   // Erhöhen des Gesammtverbrauches und des Gesamtzählers:
   // 
   "DB_Zaehler_Schicht_aktuell".Gesamt.Anzahl := "DB_Zaehler_Schicht_aktuell".Gesamt.Anzahl + 1;
   (* classic code: "DB_Zaehler_Schicht_aktuell".Gesamt.Verbrauch_K1 :=  "DB_Zaehler_Schicht_aktuell".Gesamt.Verbrauch_K1 + "DB919_ShotResultMach".ShotResult_Ma[0].Component.Comp[1].MaterialConsumption / 1000.0;*)
   "DB_Zaehler_Schicht_aktuell".Gesamt.Verbrauch_K1 :=  "DB_Zaehler_Schicht_aktuell".Gesamt.Verbrauch_K1 + "DB919_ShotResultMach".ShotResult_Ma[0].Component.Comp[1].MaterialConsumption / REAL#1000.0;
   (* classic code: "DB_Zaehler_Schicht_aktuell".Gesamt.Verbrauch_K2 :=  "DB_Zaehler_Schicht_aktuell".Gesamt.Verbrauch_K2 + "DB919_ShotResultMach".ShotResult_Ma[0].Component.Comp[2].MaterialConsumption / 1000.0;*)
   "DB_Zaehler_Schicht_aktuell".Gesamt.Verbrauch_K2 :=  "DB_Zaehler_Schicht_aktuell".Gesamt.Verbrauch_K2 + "DB919_ShotResultMach".ShotResult_Ma[0].Component.Comp[2].MaterialConsumption / REAL#1000.0;
   (* classic code: "DB_Zaehler_Schicht_aktuell".Gesamt.Verbrauch_K3 :=  "DB_Zaehler_Schicht_aktuell".Gesamt.Verbrauch_K3 + "DB919_ShotResultMach".ShotResult_Ma[0].Component.Comp[3].MaterialConsumption / 1000.0;*)
   "DB_Zaehler_Schicht_aktuell".Gesamt.Verbrauch_K3 :=  "DB_Zaehler_Schicht_aktuell".Gesamt.Verbrauch_K3 + "DB919_ShotResultMach".ShotResult_Ma[0].Component.Comp[3].MaterialConsumption / REAL#1000.0;
   (* classic code: "DB_Zaehler_Schicht_aktuell".Gesamt.Verbrauch_K4 :=  "DB_Zaehler_Schicht_aktuell".Gesamt.Verbrauch_K4 + "DB919_ShotResultMach".ShotResult_Ma[0].Component.Comp[4].MaterialConsumption / 1000.0;*)
   "DB_Zaehler_Schicht_aktuell".Gesamt.Verbrauch_K4 :=  "DB_Zaehler_Schicht_aktuell".Gesamt.Verbrauch_K4 + "DB919_ShotResultMach".ShotResult_Ma[0].Component.Comp[4].MaterialConsumption / REAL#1000.0;
   (* classic code: "DB_Zaehler_Schicht_aktuell".Gesamt.Verbrauch_K5 :=  "DB_Zaehler_Schicht_aktuell".Gesamt.Verbrauch_K5 + "DB919_ShotResultMach".ShotResult_Ma[0].Component.Comp[5].MaterialConsumption / 1000.0;*)
   "DB_Zaehler_Schicht_aktuell".Gesamt.Verbrauch_K5 :=  "DB_Zaehler_Schicht_aktuell".Gesamt.Verbrauch_K5 + "DB919_ShotResultMach".ShotResult_Ma[0].Component.Comp[5].MaterialConsumption / REAL#1000.0;
   (* classic code: "DB_Zaehler_Schicht_aktuell".Gesamt.Verbrauch_K6 :=  "DB_Zaehler_Schicht_aktuell".Gesamt.Verbrauch_K6 + "DB919_ShotResultMach".ShotResult_Ma[0].Component.Comp[6].MaterialConsumption / 1000.0;*)
   "DB_Zaehler_Schicht_aktuell".Gesamt.Verbrauch_K6 :=  "DB_Zaehler_Schicht_aktuell".Gesamt.Verbrauch_K6 + "DB919_ShotResultMach".ShotResult_Ma[0].Component.Comp[6].MaterialConsumption / REAL#1000.0;
   (* classic code: "DB_Zaehler_Schicht_aktuell".Gesamt.Verbrauch_K7 :=  "DB_Zaehler_Schicht_aktuell".Gesamt.Verbrauch_K7 + "DB919_ShotResultMach".ShotResult_Ma[0].Component.Comp[7].MaterialConsumption / 1000.0;*)
   "DB_Zaehler_Schicht_aktuell".Gesamt.Verbrauch_K7 :=  "DB_Zaehler_Schicht_aktuell".Gesamt.Verbrauch_K7 + "DB919_ShotResultMach".ShotResult_Ma[0].Component.Comp[7].MaterialConsumption / REAL#1000.0;
   (* classic code: "DB_Zaehler_Schicht_aktuell".Gesamt.Verbrauch_K8 :=  "DB_Zaehler_Schicht_aktuell".Gesamt.Verbrauch_K8 + "DB919_ShotResultMach".ShotResult_Ma[0].Component.Comp[8].MaterialConsumption / 1000.0;*)
   "DB_Zaehler_Schicht_aktuell".Gesamt.Verbrauch_K8 :=  "DB_Zaehler_Schicht_aktuell".Gesamt.Verbrauch_K8 + "DB919_ShotResultMach".ShotResult_Ma[0].Component.Comp[8].MaterialConsumption / REAL#1000.0;

   // Erhöhen des im Programm eingetragenen Schußzählers:
   // 
   // Benötigte Variablen:
   // der aktuelle Teiezähler: "DB919_ShotResultMach".ShotResult_Ma[0].General.PartID
   // 
   IF "DB919_ShotResultMach".ShotResult_Ma[0].General.PartID > 0 THEN
     #i := "DB919_ShotResultMach".ShotResult_Ma[0].General.PartID;
     "DB_Zaehler_Schicht_aktuell".Counter[#i].Anzahl := "DB_Zaehler_Schicht_aktuell".Counter[#i].Anzahl + 1;
     (* classic code: "DB_Zaehler_Schicht_aktuell".Counter[#i].Verbrauch_K1 := "DB_Zaehler_Schicht_aktuell".Counter[#i].Verbrauch_K1 + "DB919_ShotResultMach".ShotResult_Ma[0].Component.Comp[1].MaterialConsumption / 1000.0;*)
     "DB_Zaehler_Schicht_aktuell".Counter[#i].Verbrauch_K1 := "DB_Zaehler_Schicht_aktuell".Counter[#i].Verbrauch_K1 + "DB919_ShotResultMach".ShotResult_Ma[0].Component.Comp[1].MaterialConsumption / REAL#1000.0;
     (* classic code: "DB_Zaehler_Schicht_aktuell".Counter[#i].Verbrauch_K2 := "DB_Zaehler_Schicht_aktuell".Counter[#i].Verbrauch_K2 + "DB919_ShotResultMach".ShotResult_Ma[0].Component.Comp[2].MaterialConsumption / 1000.0;*)
     "DB_Zaehler_Schicht_aktuell".Counter[#i].Verbrauch_K2 := "DB_Zaehler_Schicht_aktuell".Counter[#i].Verbrauch_K2 + "DB919_ShotResultMach".ShotResult_Ma[0].Component.Comp[2].MaterialConsumption / REAL#1000.0;
     (* classic code: "DB_Zaehler_Schicht_aktuell".Counter[#i].Verbrauch_K3 := "DB_Zaehler_Schicht_aktuell".Counter[#i].Verbrauch_K3 + "DB919_ShotResultMach".ShotResult_Ma[0].Component.Comp[3].MaterialConsumption / 1000.0;*)
     "DB_Zaehler_Schicht_aktuell".Counter[#i].Verbrauch_K3 := "DB_Zaehler_Schicht_aktuell".Counter[#i].Verbrauch_K3 + "DB919_ShotResultMach".ShotResult_Ma[0].Component.Comp[3].MaterialConsumption / REAL#1000.0;
     (* classic code: "DB_Zaehler_Schicht_aktuell".Counter[#i].Verbrauch_K4 := "DB_Zaehler_Schicht_aktuell".Counter[#i].Verbrauch_K4 + "DB919_ShotResultMach".ShotResult_Ma[0].Component.Comp[4].MaterialConsumption / 1000.0;*)
     "DB_Zaehler_Schicht_aktuell".Counter[#i].Verbrauch_K4 := "DB_Zaehler_Schicht_aktuell".Counter[#i].Verbrauch_K4 + "DB919_ShotResultMach".ShotResult_Ma[0].Component.Comp[4].MaterialConsumption / REAL#1000.0;
     (* classic code: "DB_Zaehler_Schicht_aktuell".Counter[#i].Verbrauch_K5 := "DB_Zaehler_Schicht_aktuell".Counter[#i].Verbrauch_K5 + "DB919_ShotResultMach".ShotResult_Ma[0].Component.Comp[5].MaterialConsumption / 1000.0;*)
     "DB_Zaehler_Schicht_aktuell".Counter[#i].Verbrauch_K5 := "DB_Zaehler_Schicht_aktuell".Counter[#i].Verbrauch_K5 + "DB919_ShotResultMach".ShotResult_Ma[0].Component.Comp[5].MaterialConsumption / REAL#1000.0;
     (* classic code: "DB_Zaehler_Schicht_aktuell".Counter[#i].Verbrauch_K6 := "DB_Zaehler_Schicht_aktuell".Counter[#i].Verbrauch_K6 + "DB919_ShotResultMach".ShotResult_Ma[0].Component.Comp[6].MaterialConsumption / 1000.0;*)
     "DB_Zaehler_Schicht_aktuell".Counter[#i].Verbrauch_K6 := "DB_Zaehler_Schicht_aktuell".Counter[#i].Verbrauch_K6 + "DB919_ShotResultMach".ShotResult_Ma[0].Component.Comp[6].MaterialConsumption / REAL#1000.0;
     (* classic code: "DB_Zaehler_Schicht_aktuell".Counter[#i].Verbrauch_K7 := "DB_Zaehler_Schicht_aktuell".Counter[#i].Verbrauch_K7 + "DB919_ShotResultMach".ShotResult_Ma[0].Component.Comp[7].MaterialConsumption / 1000.0;*)
     "DB_Zaehler_Schicht_aktuell".Counter[#i].Verbrauch_K7 := "DB_Zaehler_Schicht_aktuell".Counter[#i].Verbrauch_K7 + "DB919_ShotResultMach".ShotResult_Ma[0].Component.Comp[7].MaterialConsumption / REAL#1000.0;
     (* classic code: "DB_Zaehler_Schicht_aktuell".Counter[#i].Verbrauch_K8 := "DB_Zaehler_Schicht_aktuell".Counter[#i].Verbrauch_K8 + "DB919_ShotResultMach".ShotResult_Ma[0].Component.Comp[8].MaterialConsumption / 1000.0;*)
     "DB_Zaehler_Schicht_aktuell".Counter[#i].Verbrauch_K8 := "DB_Zaehler_Schicht_aktuell".Counter[#i].Verbrauch_K8 + "DB919_ShotResultMach".ShotResult_Ma[0].Component.Comp[8].MaterialConsumption / REAL#1000.0;
   END_IF;
END_FUNCTION

FUNCTION "PartCounterView" : Void   // FC5002, SCL
{ S7_Optimized_Access := 'FALSE' }
VERSION : 0.1
   VAR_TEMP
      i : Int;
      CounterStartNumber : Int;
   END_VAR
BEGIN
   #CounterStartNumber := "DB_Zaehler_Anzeige".ReadWriteDeviceNo;

   IF "DB_Zaehler_Anzeige".Read THEN
     IF "DB_Zaehler_Anzeige".ViewPreShift = 0 THEN
       FOR #i := 1 TO 10 DO
         "DB_Zaehler_Anzeige".Counter[#i] :="DB_Zaehler_Schicht_aktuell".Counter[#CounterStartNumber];
         #CounterStartNumber := #CounterStartNumber +1;
       END_FOR;
       "DB_Zaehler_Anzeige".Gesamt := "DB_Zaehler_Schicht_aktuell".Gesamt;
       "DB_Zaehler_Anzeige".MH_Counter_ActualShift := "DB_Zaehler_Schicht_aktuell".MH_Counter;
     ELSE
       FOR #i := 1 TO 10 DO
         "DB_Zaehler_Anzeige".Counter[#i] :="DB_Zaehler_Schicht_Vorherige".Counter[#CounterStartNumber];
         #CounterStartNumber := #CounterStartNumber +1;
       END_FOR;
       "DB_Zaehler_Anzeige".Gesamt := "DB_Zaehler_Schicht_Vorherige".Gesamt;
       "DB_Zaehler_Anzeige".MH_Counter_ActualShift := "DB_Zaehler_Schicht_Vorherige".MH_Counter;
     END_IF;

     FOR #i := 1 TO 16 DO
       "DB_Zaehler_Anzeige".MH_Counter_ActualShift[#i] := "DB_Zaehler_Schicht_aktuell".MH_Counter[#i];
       "DB_Zaehler_Anzeige".MH_Counter_PreShift[#i] :=  "DB_Zaehler_Schicht_Vorherige".MH_Counter[#i];
     END_FOR;

   END_IF;

   "DB_Zaehler_Anzeige".Read := false;
END_FUNCTION

FUNCTION "PartCounterCopy" : Void   // FC5003, SCL
{ S7_Optimized_Access := 'FALSE' }
VERSION : 0.1
   VAR_TEMP
      i : Int;
   END_VAR
BEGIN
   // 
   // Shift the part counter at the begining of a new shift!
   // 
   "DB_Zaehler_Schicht_Vorherige".Gesamt := "DB_Zaehler_Schicht_aktuell".Gesamt;
   "DB_Zaehler_Schicht_Vorherige".Counter := "DB_Zaehler_Schicht_aktuell".Counter;
   "DB_Zaehler_Schicht_Vorherige".MH_Counter := "DB_Zaehler_Schicht_aktuell".MH_Counter;

   // Reset the amount of Counts and weight
   // 
   "DB_Zaehler_Schicht_aktuell".Gesamt.Anzahl := 0;
   (* classic code: "DB_Zaehler_Schicht_aktuell".Gesamt.Verbrauch_K1 := 0.0;*)
   "DB_Zaehler_Schicht_aktuell".Gesamt.Verbrauch_K1 := REAL#0.0;
   (* classic code: "DB_Zaehler_Schicht_aktuell".Gesamt.Verbrauch_K2 := 0.0;*)
   "DB_Zaehler_Schicht_aktuell".Gesamt.Verbrauch_K2 := REAL#0.0;
   (* classic code: "DB_Zaehler_Schicht_aktuell".Gesamt.Verbrauch_K3 := 0.0;*)
   "DB_Zaehler_Schicht_aktuell".Gesamt.Verbrauch_K3 := REAL#0.0;
   (* classic code: "DB_Zaehler_Schicht_aktuell".Gesamt.Verbrauch_K4 := 0.0;*)
   "DB_Zaehler_Schicht_aktuell".Gesamt.Verbrauch_K4 := REAL#0.0;
   (* classic code: "DB_Zaehler_Schicht_aktuell".Gesamt.Verbrauch_K5 := 0.0;*)
   "DB_Zaehler_Schicht_aktuell".Gesamt.Verbrauch_K5 := REAL#0.0;
   (* classic code: "DB_Zaehler_Schicht_aktuell".Gesamt.Verbrauch_K6 := 0.0;*)
   "DB_Zaehler_Schicht_aktuell".Gesamt.Verbrauch_K6 := REAL#0.0;
   (* classic code: "DB_Zaehler_Schicht_aktuell".Gesamt.Verbrauch_K7 := 0.0;*)
   "DB_Zaehler_Schicht_aktuell".Gesamt.Verbrauch_K7 := REAL#0.0;
   (* classic code: "DB_Zaehler_Schicht_aktuell".Gesamt.Verbrauch_K8 := 0.0;*)
   "DB_Zaehler_Schicht_aktuell".Gesamt.Verbrauch_K8 := REAL#0.0;

   FOR #i := 1 TO 120 DO
     "DB_Zaehler_Schicht_aktuell".Counter[#i].Anzahl := 0;
     (* classic code: "DB_Zaehler_Schicht_aktuell".Counter[#i].Verbrauch_K1 := 0.0;*)
     "DB_Zaehler_Schicht_aktuell".Counter[#i].Verbrauch_K1 := REAL#0.0;
     (* classic code: "DB_Zaehler_Schicht_aktuell".Counter[#i].Verbrauch_K2 := 0.0;*)
     "DB_Zaehler_Schicht_aktuell".Counter[#i].Verbrauch_K2 := REAL#0.0;
     (* classic code: "DB_Zaehler_Schicht_aktuell".Counter[#i].Verbrauch_K3 := 0.0;*)
     "DB_Zaehler_Schicht_aktuell".Counter[#i].Verbrauch_K3 := REAL#0.0;
     (* classic code: "DB_Zaehler_Schicht_aktuell".Counter[#i].Verbrauch_K4 := 0.0;*)
     "DB_Zaehler_Schicht_aktuell".Counter[#i].Verbrauch_K4 := REAL#0.0;
     (* classic code: "DB_Zaehler_Schicht_aktuell".Counter[#i].Verbrauch_K5 := 0.0;*)
     "DB_Zaehler_Schicht_aktuell".Counter[#i].Verbrauch_K5 := REAL#0.0;
     (* classic code: "DB_Zaehler_Schicht_aktuell".Counter[#i].Verbrauch_K6 := 0.0;*)
     "DB_Zaehler_Schicht_aktuell".Counter[#i].Verbrauch_K6 := REAL#0.0;
     (* classic code: "DB_Zaehler_Schicht_aktuell".Counter[#i].Verbrauch_K7 := 0.0;*)
     "DB_Zaehler_Schicht_aktuell".Counter[#i].Verbrauch_K7 := REAL#0.0;
     (* classic code: "DB_Zaehler_Schicht_aktuell".Counter[#i].Verbrauch_K8 := 0.0;*)
     "DB_Zaehler_Schicht_aktuell".Counter[#i].Verbrauch_K8 := REAL#0.0;
     (* classic code: "DB_Zaehler_Schicht_aktuell".Counter[#i].Verbrauch_K8 := 0.0;*)
     "DB_Zaehler_Schicht_aktuell".Counter[#i].Verbrauch_K8 := REAL#0.0;
   END_FOR;

   FOR #i := 1 TO 16 DO
     "DB_Zaehler_Schicht_aktuell".MH_Counter[#i] := 0;
   END_FOR;

   "DB_Zaehler_Anzeige".Schichtwechsel := 0;
END_FUNCTION

FUNCTION "FC5011_InterfaceHydraulik" : Void   // FC5011, SCL
{ S7_Optimized_Access := 'FALSE' }
VERSION : 0.1
   VAR_INPUT
      Enable : Bool;
   END_VAR
BEGIN
   // Status: DB612_Hydraulic_State
   // Values: DB721_MH_Hydraulic
   // Faults: DB821_Error_Hydraulic
   // 

   // Read the Values only once after open the window or change the Number
   // 
   IF ("DB611_Hydraulic_State".ReadDeviceNo <> "DB611_Hydraulic_State".ActualDeviceNo) OR "DB611_Hydraulic_State".Read THEN
       "DB611_Hydraulic_State".ActualDeviceNo := "DB611_Hydraulic_State".ReadDeviceNo;

       // Status
       "DB611_Hydraulic_State".MH_Hydraulic[0] := "DB611_Hydraulic_State".MH_Hydraulic["DB611_Hydraulic_State".ReadDeviceNo];
       "DB611_Hydraulic_State".S_Hydraulic[0] := "DB611_Hydraulic_State".S_Hydraulic["DB611_Hydraulic_State".ReadDeviceNo];
       "DB611_Hydraulic_State".NZL_Hydraulic[0] := "DB611_Hydraulic_State".NZL_Hydraulic["DB611_Hydraulic_State".ReadDeviceNo];
       // Setvalues 
       "DB721_MH_Hydraulic".Option[0] := "DB721_MH_Hydraulic".Option["DB611_Hydraulic_State".ReadDeviceNo];
       "DB721_MH_Hydraulic".MH_Hyd[0] := "DB721_MH_Hydraulic".MH_Hyd["DB611_Hydraulic_State".ReadDeviceNo];
       "DB721_MH_Hydraulic".S_Hyd[0] := "DB721_MH_Hydraulic".S_Hyd["DB611_Hydraulic_State".ReadDeviceNo];
       "DB721_MH_Hydraulic".NZL_Hyd[0] := "DB721_MH_Hydraulic".NZL_Hyd["DB611_Hydraulic_State".ReadDeviceNo];

       "DB611_Hydraulic_State".Read := FALSE;

   END_IF;

   // If not the hydraulic page was selectet don't copy the values   
   IF "TP-Bereichszeiger".Picturenumber.Bildnummer = 2 THEN
   // If a status changed by operator copy this to the select number and do not read all status values
       IF "DB611_Hydraulic_State".MH_Hydraulic["DB611_Hydraulic_State".ReadDeviceNo].Switch_Hydraulic_ON_OFF <> "DB611_Hydraulic_State".MH_Hydraulic[0].Switch_Hydraulic_ON_OFF OR
           "DB611_Hydraulic_State".S_Hydraulic["DB611_Hydraulic_State".ReadDeviceNo].Switch_Hydraulic_ON_OFF <> "DB611_Hydraulic_State".S_Hydraulic[0].Switch_Hydraulic_ON_OFF OR
           "DB611_Hydraulic_State".NZL_Hydraulic["DB611_Hydraulic_State".ReadDeviceNo].Switch_Hydraulic_ON_OFF <> "DB611_Hydraulic_State".NZL_Hydraulic[0].Switch_Hydraulic_ON_OFF
       THEN
           // copy the [0] switch to the selected switch
           "DB611_Hydraulic_State".MH_Hydraulic["DB611_Hydraulic_State".ReadDeviceNo].Switch_Hydraulic_ON_OFF := "DB611_Hydraulic_State".MH_Hydraulic[0].Switch_Hydraulic_ON_OFF;
           "DB611_Hydraulic_State".S_Hydraulic["DB611_Hydraulic_State".ReadDeviceNo].Switch_Hydraulic_ON_OFF := "DB611_Hydraulic_State".S_Hydraulic[0].Switch_Hydraulic_ON_OFF;
           "DB611_Hydraulic_State".NZL_Hydraulic["DB611_Hydraulic_State".ReadDeviceNo].Switch_Hydraulic_ON_OFF := "DB611_Hydraulic_State".NZL_Hydraulic[0].Switch_Hydraulic_ON_OFF;
       ELSE
           // Read the status of the selected hydraulic
           "DB611_Hydraulic_State".MH_Hydraulic[0] := "DB611_Hydraulic_State".MH_Hydraulic["DB611_Hydraulic_State".ReadDeviceNo];
           "DB611_Hydraulic_State".S_Hydraulic[0] :="DB611_Hydraulic_State".S_Hydraulic["DB611_Hydraulic_State".ReadDeviceNo];
           "DB611_Hydraulic_State".NZL_Hydraulic[0] := "DB611_Hydraulic_State".NZL_Hydraulic["DB611_Hydraulic_State".ReadDeviceNo];
       END_IF;

   END_IF;

   // Write the values 
   IF "DB611_Hydraulic_State".Write = TRUE THEN

       // Values 
       "DB721_MH_Hydraulic".Option["DB611_Hydraulic_State".ReadDeviceNo] := "DB721_MH_Hydraulic".Option[0];
       "DB721_MH_Hydraulic".MH_Hyd["DB611_Hydraulic_State".ReadDeviceNo] := "DB721_MH_Hydraulic".MH_Hyd[0];
       "DB721_MH_Hydraulic".S_Hyd["DB611_Hydraulic_State".ReadDeviceNo] := "DB721_MH_Hydraulic".S_Hyd[0];
       "DB721_MH_Hydraulic".NZL_Hyd["DB611_Hydraulic_State".ReadDeviceNo] := "DB721_MH_Hydraulic".NZL_Hyd[0];

       "DB611_Hydraulic_State".Write := FALSE;

   END_IF;

   // Show the actual values every time:
   "DB611_Hydraulic_State".MH_Hydraulic[0].HourCounter := "DB611_Hydraulic_State".MH_Hydraulic["DB611_Hydraulic_State".ReadDeviceNo].HourCounter;
   // Show the actual faults every time
   "DB821_Error_Hydraulic".MH_Hydraulic[0] := "DB821_Error_Hydraulic".MH_Hydraulic["DB611_Hydraulic_State".ReadDeviceNo];
   "DB821_Error_Hydraulic".S_Hydraulic[0] := "DB821_Error_Hydraulic".S_Hydraulic["DB611_Hydraulic_State".ReadDeviceNo];
   "DB821_Error_Hydraulic".NZL_Hydraulic[0] := "DB821_Error_Hydraulic".NZL_Hydraulic["DB611_Hydraulic_State".ReadDeviceNo];
END_FUNCTION

FUNCTION "FC5012_InterfaceTank" : Void   // FC5012, SCL
{ S7_Optimized_Access := 'FALSE' }
VERSION : 0.1
   VAR_INPUT
      Enable : Bool;
   END_VAR
BEGIN
   // Status: DB612_Tank_State
   // Values: DB602_PV_Tank
   // Config: DB702_Tank_Value
   // Faults: DB822_Error_Tank
   // 

   // Read the Values only once after open the window or change the Number
   // 
   IF ("DB612_Tank_State".ReadDeviceNo <> "DB612_Tank_State".ActualDeviceNo) OR "DB612_Tank_State".Read THEN
       "DB612_Tank_State".ActualDeviceNo := "DB612_Tank_State".ReadDeviceNo;

       // Setvalues 
       "DB602_PV_Tank".Tank[0] := "DB602_PV_Tank".Tank["DB612_Tank_State".ReadDeviceNo];
       // Status
       "DB612_Tank_State".Tank[0] := "DB612_Tank_State".Tank["DB612_Tank_State".ReadDeviceNo];
       "DB612_Tank_State".Agitator[0] := "DB612_Tank_State".Agitator["DB612_Tank_State".ReadDeviceNo];
       "DB612_Tank_State".Vacuum[0] := "DB612_Tank_State".Vacuum["DB612_Tank_State".ReadDeviceNo];
       "DB612_Tank_State".AgitatorBarell[0] := "DB612_Tank_State".AgitatorBarell["DB612_Tank_State".ReadDeviceNo];
       "DB612_Tank_State".ControllerTankTemp[0] := "DB612_Tank_State".ControllerTankTemp["DB612_Tank_State".ReadDeviceNo];
       "DB612_Tank_State".ControllerTankJacketHeater[0] := "DB612_Tank_State".ControllerTankJacketHeater["DB612_Tank_State".ReadDeviceNo];
       "DB612_Tank_State".CirculationPump[0] := "DB612_Tank_State".CirculationPump["DB612_Tank_State".ReadDeviceNo];
       // Config values
       "DB702_Tank_Value".Tank[0] := "DB702_Tank_Value".Tank["DB612_Tank_State".ReadDeviceNo];
       "DB702_Tank_Value".AgitatorBarell[0] := "DB702_Tank_Value".AgitatorBarell["DB612_Tank_State".ReadDeviceNo];
       "DB702_Tank_Value".Pt2_Controller[0] := "DB702_Tank_Value".Pt2_Controller["DB612_Tank_State".ReadDeviceNo];
       "DB702_Tank_Value".Pt2_ControllerBarell[0] := "DB702_Tank_Value".Pt2_ControllerBarell["DB612_Tank_State".ReadDeviceNo];
       "DB702_Tank_Value".CirculationPump[0] := "DB702_Tank_Value".CirculationPump["DB612_Tank_State".ReadDeviceNo];

       "DB612_Tank_State".Read := FALSE;

   END_IF;

   // If not the Tank page was selectet don't copy the values   
   IF "TP-Bereichszeiger".Picturenumber.Bildnummer = 6 THEN
     // If a status changed by operator copy this to the select number and do not read all status values
       IF "DB612_Tank_State".Tank["DB612_Tank_State".ReadDeviceNo].Switch_Refilling_ON_OFF <> "DB612_Tank_State".Tank[0].Switch_Refilling_ON_OFF OR
           "DB612_Tank_State".Tank["DB612_Tank_State".ReadDeviceNo].ButtonLeakageMonitorOFF <> "DB612_Tank_State".Tank[0].ButtonLeakageMonitorOFF OR
           "DB612_Tank_State".Agitator["DB612_Tank_State".ReadDeviceNo].Switch_Drive_ON_OFF <> "DB612_Tank_State".Agitator[0].Switch_Drive_ON_OFF OR
           "DB612_Tank_State".Vacuum["DB612_Tank_State".ReadDeviceNo].Switch_Vacuum_ON_OFF <> "DB612_Tank_State".Vacuum[0].Switch_Vacuum_ON_OFF OR
           "DB612_Tank_State".AgitatorBarell["DB612_Tank_State".ReadDeviceNo].Switch_Drive_ON_OFF <> "DB612_Tank_State".AgitatorBarell[0].Switch_Drive_ON_OFF OR
           "DB612_Tank_State".ControllerTankTemp["DB612_Tank_State".ReadDeviceNo].Switch_Temp_ON_OFF <> "DB612_Tank_State".ControllerTankTemp[0].Switch_Temp_ON_OFF OR
           "DB612_Tank_State".ControllerTankJacketHeater["DB612_Tank_State".ReadDeviceNo].Switch_Temp_ON_OFF <> "DB612_Tank_State".ControllerTankJacketHeater[0].Switch_Temp_ON_OFF OR
           "DB612_Tank_State".CirculationPump["DB612_Tank_State".ReadDeviceNo].Switch_Drive_ON_OFF <> "DB612_Tank_State".CirculationPump[0].Switch_Drive_ON_OFF OR
           "DB612_Tank_State".Tank["DB612_Tank_State".ReadDeviceNo].Switch_Refilling_from_Barrel_ON_OFF <> "DB612_Tank_State".Tank[0].Switch_Refilling_from_Barrel_ON_OFF
       THEN
           // copy the [0] switch to the selected switch
           "DB612_Tank_State".Tank["DB612_Tank_State".ReadDeviceNo].Switch_Refilling_ON_OFF := "DB612_Tank_State".Tank[0].Switch_Refilling_ON_OFF;
           "DB612_Tank_State".Tank["DB612_Tank_State".ReadDeviceNo].ButtonLeakageMonitorOFF := "DB612_Tank_State".Tank[0].ButtonLeakageMonitorOFF;
           "DB612_Tank_State".Agitator["DB612_Tank_State".ReadDeviceNo].Switch_Drive_ON_OFF := "DB612_Tank_State".Agitator[0].Switch_Drive_ON_OFF;
           "DB612_Tank_State".Vacuum["DB612_Tank_State".ReadDeviceNo].Switch_Vacuum_ON_OFF := "DB612_Tank_State".Vacuum[0].Switch_Vacuum_ON_OFF;
           "DB612_Tank_State".AgitatorBarell["DB612_Tank_State".ReadDeviceNo].Switch_Drive_ON_OFF := "DB612_Tank_State".AgitatorBarell[0].Switch_Drive_ON_OFF;
           "DB612_Tank_State".ControllerTankTemp["DB612_Tank_State".ReadDeviceNo].Switch_Temp_ON_OFF := "DB612_Tank_State".ControllerTankTemp[0].Switch_Temp_ON_OFF;
           "DB612_Tank_State".ControllerTankJacketHeater["DB612_Tank_State".ReadDeviceNo].Switch_Temp_ON_OFF := "DB612_Tank_State".ControllerTankJacketHeater[0].Switch_Temp_ON_OFF;
           "DB612_Tank_State".CirculationPump["DB612_Tank_State".ReadDeviceNo].Switch_Drive_ON_OFF := "DB612_Tank_State".CirculationPump[0].Switch_Drive_ON_OFF;
           "DB612_Tank_State".Tank["DB612_Tank_State".ReadDeviceNo].Switch_Refilling_from_Barrel_ON_OFF := "DB612_Tank_State".Tank[0].Switch_Refilling_from_Barrel_ON_OFF;
       ELSE
           // Read the status of the selected hydraulic
           "DB612_Tank_State".Tank[0] := "DB612_Tank_State".Tank["DB612_Tank_State".ReadDeviceNo];
           "DB612_Tank_State".Agitator[0] := "DB612_Tank_State".Agitator["DB612_Tank_State".ReadDeviceNo];
           "DB612_Tank_State".Vacuum[0] := "DB612_Tank_State".Vacuum["DB612_Tank_State".ReadDeviceNo];
           "DB612_Tank_State".AgitatorBarell[0] := "DB612_Tank_State".AgitatorBarell["DB612_Tank_State".ReadDeviceNo];
           "DB612_Tank_State".ControllerTankTemp[0] := "DB612_Tank_State".ControllerTankTemp["DB612_Tank_State".ReadDeviceNo];
           "DB612_Tank_State".ControllerTankJacketHeater[0] := "DB612_Tank_State".ControllerTankJacketHeater["DB612_Tank_State".ReadDeviceNo];
           "DB612_Tank_State".CirculationPump[0] := "DB612_Tank_State".CirculationPump["DB612_Tank_State".ReadDeviceNo];

           "DB905_GWK".State[0].Act_value_tempering_unit := "DB905_GWK".State["DB612_Tank_State".ReadDeviceNo].Act_value_tempering_unit;
           "DB905_GWK".State[0].Fault_state := "DB905_GWK".State["DB612_Tank_State".ReadDeviceNo].Fault_state;
       END_IF;

   END_IF;

   // Write the request for the switches once
   IF "DB612_Tank_State".Write = TRUE OR "DB702_Tank_Value".Write = TRUE THEN
       // Values 
       "DB602_PV_Tank".Tank["DB612_Tank_State".ReadDeviceNo] := "DB602_PV_Tank".Tank[0];
       "DB702_Tank_Value".Tank["DB612_Tank_State".ReadDeviceNo] := "DB702_Tank_Value".Tank[0];
       "DB702_Tank_Value".AgitatorBarell["DB612_Tank_State".ReadDeviceNo] := "DB702_Tank_Value".AgitatorBarell[0];
       "DB702_Tank_Value".Pt2_Controller["DB612_Tank_State".ReadDeviceNo] := "DB702_Tank_Value".Pt2_Controller[0];
       "DB702_Tank_Value".Pt2_ControllerBarell["DB612_Tank_State".ReadDeviceNo] := "DB702_Tank_Value".Pt2_ControllerBarell[0];
       "DB702_Tank_Value".CirculationPump["DB612_Tank_State".ReadDeviceNo] := "DB702_Tank_Value".CirculationPump[0];

       // Config Bits schieben
       "DB702_Tank_Value".Tank[0].Agitator.Config_bit_Converter := "DB702_Tank_Value".Tank[0].With_Agitator_Converter;
       "DB702_Tank_Value".Tank["DB612_Tank_State".ReadDeviceNo].Agitator.Config_bit_Converter := "DB702_Tank_Value".Tank[0].Agitator.Config_bit_Converter;


       "DB612_Tank_State".Write := FALSE;
       "DB702_Tank_Value".Write := FALSE;

   END_IF;

   // Show the actual faults every time
   "DB822_Error_Tank".FeedPump[0] := "DB822_Error_Tank".FeedPump["DB612_Tank_State".ReadDeviceNo];
   "DB822_Error_Tank".Agitator[0] := "DB822_Error_Tank".Agitator["DB612_Tank_State".ReadDeviceNo];
   "DB822_Error_Tank".Refilling_Tank[0] := "DB822_Error_Tank".Refilling_Tank["DB612_Tank_State".ReadDeviceNo];
   "DB822_Error_Tank".CirculationPump[0] := "DB822_Error_Tank".CirculationPump["DB612_Tank_State".ReadDeviceNo];
   "DB822_Error_Tank".RefillingStation[0] := "DB822_Error_Tank".RefillingStation["DB612_Tank_State".ReadDeviceNo];
   "DB822_Error_Tank".Temperature_Heatexchange[0] := "DB822_Error_Tank".Temperature_Heatexchange["DB612_Tank_State".ReadDeviceNo];
   "DB822_Error_Tank".ControllerTankTemp[0] := "DB822_Error_Tank".ControllerTankTemp["DB612_Tank_State".ReadDeviceNo];
   "DB822_Error_Tank".ControllerTankJacketHeater[0] := "DB822_Error_Tank".ControllerTankJacketHeater["DB612_Tank_State".ReadDeviceNo];
   "DB822_Error_Tank".ControllerBarellTemp[0] := "DB822_Error_Tank".ControllerBarellTemp["DB612_Tank_State".ReadDeviceNo];
   "DB822_Error_Tank".Vacuum[0] := "DB822_Error_Tank".Vacuum["DB612_Tank_State".ReadDeviceNo];
   "DB822_Error_Tank".CoverLift[0] := "DB822_Error_Tank".CoverLift["DB612_Tank_State".ReadDeviceNo];
   "DB822_Error_Tank".LevelRefillingStation[0] := "DB822_Error_Tank".LevelRefillingStation["DB612_Tank_State".ReadDeviceNo];
   "DB822_Error_Tank".TempRefillingStation[0] := "DB822_Error_Tank".TempRefillingStation["DB612_Tank_State".ReadDeviceNo];
   "DB822_Error_Tank".LeakageMonitor[0] := "DB822_Error_Tank".LeakageMonitor["DB612_Tank_State".ReadDeviceNo];
   "DB822_Error_Tank".AgitatorBarrel[0] := "DB822_Error_Tank".AgitatorBarrel["DB612_Tank_State".ReadDeviceNo];
   "DB822_Error_Tank".Pentan[0] := "DB822_Error_Tank".Pentan["DB612_Tank_State".ReadDeviceNo];
END_FUNCTION

FUNCTION "FC5013_InterfaceMetering" : Void   // FC5013, SCL
{ S7_Optimized_Access := 'FALSE' }
VERSION : 0.1
   VAR_INPUT
      Enable : Bool;
   END_VAR
BEGIN

   // When the selected number change or the read bit was set 
   // read the set values once
   IF ("DB613_Komponent_State".ReadDeviceNo <> "DB613_Komponent_State".ActualDeviceNo) OR "DB613_Komponent_State".Read THEN
       "DB613_Komponent_State".ActualDeviceNo := "DB613_Komponent_State".ReadDeviceNo;

       // Read all prozess values for the component plunger
       "DB601_PV_Plunger".Component[0] := "DB601_PV_Plunger".Component["DB613_Komponent_State".ReadDeviceNo];
       // Read all prozess values
       "DB608_PV_Metering".Metering[0].Pressure := "DB608_PV_Metering".Metering["DB613_Komponent_State".ReadDeviceNo].Pressure;
       "DB608_PV_Metering".Metering[0].Flow := "DB608_PV_Metering".Metering["DB613_Komponent_State".ReadDeviceNo].Flow;
       "DB608_PV_Metering".Metering[0].Temperature := "DB608_PV_Metering".Metering["DB613_Komponent_State".ReadDeviceNo].Temperature;
       "DB608_PV_Metering".Metering[0].Pre_Pressure := "DB608_PV_Metering".Metering["DB613_Komponent_State".ReadDeviceNo].Pre_Pressure;
       "DB608_PV_Metering".Metering[0].MixingRatio := "DB608_PV_Metering".Metering["DB613_Komponent_State".ReadDeviceNo].MixingRatio;
       "DB608_PV_Metering".HeatexchangerHP[0] := "DB608_PV_Metering".HeatexchangerHP["DB613_Komponent_State".ReadDeviceNo];
       "DB608_PV_Metering".HeatexchangerLP[0] := "DB608_PV_Metering".HeatexchangerLP["DB613_Komponent_State".ReadDeviceNo];
       "DB608_PV_Metering".Heating[0] := "DB608_PV_Metering".Heating["DB613_Komponent_State".ReadDeviceNo];

       // Status
       "DB613_Komponent_State".FeedPump[0] := "DB613_Komponent_State".FeedPump["DB613_Komponent_State".ReadDeviceNo];
       "DB613_Komponent_State".EdgeFilter[0] := "DB613_Komponent_State".EdgeFilter["DB613_Komponent_State".ReadDeviceNo];
       "DB613_Komponent_State".MeteringPump[0] := "DB613_Komponent_State".MeteringPump["DB613_Komponent_State".ReadDeviceNo];
       "DB613_Komponent_State".Cylinder[0] := "DB613_Komponent_State".Cylinder["DB613_Komponent_State".ReadDeviceNo];
       "DB613_Komponent_State".FlowPumpMin[0] := "DB613_Komponent_State".FlowPumpMin["DB613_Komponent_State".ReadDeviceNo];
       "DB613_Komponent_State".FlowPumpMax[0] := "DB613_Komponent_State".FlowPumpMax["DB613_Komponent_State".ReadDeviceNo];
       "DB613_Komponent_State".FlowPump[0] := "DB613_Komponent_State".FlowPump["DB613_Komponent_State".ReadDeviceNo];
       "DB613_Komponent_State".FlowPumpQPB[0] := "DB613_Komponent_State".FlowPumpQPB["DB613_Komponent_State".ReadDeviceNo];
       "DB613_Komponent_State".PressurePumpQPB[0] := "DB613_Komponent_State".PressurePumpQPB["DB613_Komponent_State".ReadDeviceNo];
       "DB613_Komponent_State".FlowPumpPContr[0] := "DB613_Komponent_State".FlowPumpPContr["DB613_Komponent_State".ReadDeviceNo];
       "DB613_Komponent_State".AbortComponent[0] := "DB613_Komponent_State".AbortComponent["DB613_Komponent_State".ReadDeviceNo];
       "DB613_Komponent_State".ServoECylinder[0] := "DB613_Komponent_State".ServoECylinder["DB613_Komponent_State".ReadDeviceNo];
       "DB613_Komponent_State".GroupStatus[0] := "DB613_Komponent_State".GroupStatus["DB613_Komponent_State".ReadDeviceNo];
       "DB613_Komponent_State".HeatexchangerHP[0] := "DB613_Komponent_State".HeatexchangerHP["DB613_Komponent_State".ReadDeviceNo];
       "DB613_Komponent_State".HeatexchangerLP[0] := "DB613_Komponent_State".HeatexchangerLP["DB613_Komponent_State".ReadDeviceNo];
       "DB613_Komponent_State".Heating[0] := "DB613_Komponent_State".Heating["DB613_Komponent_State".ReadDeviceNo];

       // Read all values for the auxilary drives
       "DB751_auxiliaryDriveMetering".FeedingPump[0] := "DB751_auxiliaryDriveMetering".FeedingPump["DB613_Komponent_State".ReadDeviceNo];
       "DB751_auxiliaryDriveMetering".EdgeFilter[0] := "DB751_auxiliaryDriveMetering".EdgeFilter["DB613_Komponent_State".ReadDeviceNo];
       "DB751_auxiliaryDriveMetering".HeatConverter[0] := "DB751_auxiliaryDriveMetering".HeatConverter["DB613_Komponent_State".ReadDeviceNo];
       "DB751_auxiliaryDriveMetering".HeatexchangerHP[0] := "DB751_auxiliaryDriveMetering".HeatexchangerHP["DB613_Komponent_State".ReadDeviceNo];
       "DB751_auxiliaryDriveMetering".HeatexchangerLP[0] := "DB751_auxiliaryDriveMetering".HeatexchangerLP["DB613_Komponent_State".ReadDeviceNo];
       "DB751_auxiliaryDriveMetering".FeedingPumpControler[0] := "DB751_auxiliaryDriveMetering".FeedingPumpControler["DB613_Komponent_State".ReadDeviceNo];

       // Read all values for the component pumps
       "DB753_MeteringPump".HeatingController[0] := "DB753_MeteringPump".HeatingController["DB613_Komponent_State".ReadDeviceNo];
       "DB753_MeteringPump".Heating[0] := "DB753_MeteringPump".Heating["DB613_Komponent_State".ReadDeviceNo];
       "DB753_MeteringPump".Pump[0] := "DB753_MeteringPump".Pump["DB613_Komponent_State".ReadDeviceNo];

       // Read all values for the component plunger
       "DB762_Cylinder".Cylinder[0] := "DB762_Cylinder".Cylinder["DB613_Komponent_State".ReadDeviceNo];

       // Read special Flow values 
       "DB902_ConfFlow_PV".Flow[0].controltime := "DB902_ConfFlow_PV".Flow["DB613_Komponent_State".ReadDeviceNo].controltime;

       "DB613_Komponent_State".Read := FALSE;

   END_IF;

   // If not the component page was selectet don't copy the values   
   IF "TP-Bereichszeiger".Picturenumber.Bildnummer = 10 THEN
       // If a status changed by operator copy this to the select number and do not read all status values
       IF     "DB613_Komponent_State".FeedPump["DB613_Komponent_State".ReadDeviceNo].Switch_Drive_ON_OFF <> "DB613_Komponent_State".FeedPump[0].Switch_Drive_ON_OFF OR
           "DB613_Komponent_State".EdgeFilter["DB613_Komponent_State".ReadDeviceNo].Switch_Drive_ON_OFF <> "DB613_Komponent_State".EdgeFilter[0].Switch_Drive_ON_OFF OR
           "DB613_Komponent_State".AbortComponent["DB613_Komponent_State".ReadDeviceNo].Abort_ON_OFF <> "DB613_Komponent_State".AbortComponent[0].Abort_ON_OFF OR
           "DB613_Komponent_State".HeatexchangerHP["DB613_Komponent_State".ReadDeviceNo].Switch_Temp_ON_OFF <> "DB613_Komponent_State".HeatexchangerHP[0].Switch_Temp_ON_OFF OR
           "DB613_Komponent_State".HeatexchangerLP["DB613_Komponent_State".ReadDeviceNo].Switch_Temp_ON_OFF <> "DB613_Komponent_State".HeatexchangerLP[0].Switch_Temp_ON_OFF
       THEN
           // copy the [0] switch to the selected switch
           "DB613_Komponent_State".FeedPump["DB613_Komponent_State".ReadDeviceNo].Switch_Drive_ON_OFF := "DB613_Komponent_State".FeedPump[0].Switch_Drive_ON_OFF;
           "DB613_Komponent_State".EdgeFilter["DB613_Komponent_State".ReadDeviceNo].Switch_Drive_ON_OFF := "DB613_Komponent_State".EdgeFilter[0].Switch_Drive_ON_OFF;
           "DB613_Komponent_State".AbortComponent["DB613_Komponent_State".ReadDeviceNo].Abort_ON_OFF := "DB613_Komponent_State".AbortComponent[0].Abort_ON_OFF;
           "DB613_Komponent_State".HeatexchangerHP["DB613_Komponent_State".ReadDeviceNo].Switch_Temp_ON_OFF := "DB613_Komponent_State".HeatexchangerHP[0].Switch_Temp_ON_OFF;
           "DB613_Komponent_State".HeatexchangerLP["DB613_Komponent_State".ReadDeviceNo].Switch_Temp_ON_OFF := "DB613_Komponent_State".HeatexchangerLP[0].Switch_Temp_ON_OFF;
       ELSE
           // Read the status of the selected hydraulic
           "DB613_Komponent_State".FeedPump[0] := "DB613_Komponent_State".FeedPump["DB613_Komponent_State".ReadDeviceNo];
           "DB613_Komponent_State".EdgeFilter[0] := "DB613_Komponent_State".EdgeFilter["DB613_Komponent_State".ReadDeviceNo];
           "DB613_Komponent_State".MeteringPump[0] := "DB613_Komponent_State".MeteringPump["DB613_Komponent_State".ReadDeviceNo];
           "DB613_Komponent_State".Cylinder[0] := "DB613_Komponent_State".Cylinder["DB613_Komponent_State".ReadDeviceNo];
           "DB613_Komponent_State".FlowPumpMin[0] := "DB613_Komponent_State".FlowPumpMin["DB613_Komponent_State".ReadDeviceNo];
           "DB613_Komponent_State".FlowPumpMax[0] := "DB613_Komponent_State".FlowPumpMax["DB613_Komponent_State".ReadDeviceNo];
           "DB613_Komponent_State".FlowPump[0] := "DB613_Komponent_State".FlowPump["DB613_Komponent_State".ReadDeviceNo];
           "DB613_Komponent_State".FlowPumpQPB[0] := "DB613_Komponent_State".FlowPumpQPB["DB613_Komponent_State".ReadDeviceNo];
           "DB613_Komponent_State".PressurePumpQPB[0] := "DB613_Komponent_State".PressurePumpQPB["DB613_Komponent_State".ReadDeviceNo];
           "DB613_Komponent_State".FlowPumpPContr[0] := "DB613_Komponent_State".FlowPumpPContr["DB613_Komponent_State".ReadDeviceNo];
           "DB613_Komponent_State".AbortComponent[0] := "DB613_Komponent_State".AbortComponent["DB613_Komponent_State".ReadDeviceNo];
           "DB613_Komponent_State".ServoECylinder[0] := "DB613_Komponent_State".ServoECylinder["DB613_Komponent_State".ReadDeviceNo];
           "DB613_Komponent_State".GroupStatus[0] := "DB613_Komponent_State".GroupStatus["DB613_Komponent_State".ReadDeviceNo];
           "DB613_Komponent_State".HeatexchangerHP[0] := "DB613_Komponent_State".HeatexchangerHP["DB613_Komponent_State".ReadDeviceNo];
           "DB613_Komponent_State".HeatexchangerLP[0] := "DB613_Komponent_State".HeatexchangerLP["DB613_Komponent_State".ReadDeviceNo];
       END_IF;

   END_IF;

   // If not the component heating page was selectet don't copy the values   
   IF "TP-Bereichszeiger".Picturenumber.Bildnummer = 39 THEN
       // If a status changed by operator copy this to the select number and do not read all status values
       IF     "DB613_Komponent_State".Heating["DB613_Komponent_State".ReadDeviceNo].Heating[1].Switch_ON_OFF <> "DB613_Komponent_State".Heating[0].Heating[1].Switch_ON_OFF OR
           "DB613_Komponent_State".Heating["DB613_Komponent_State".ReadDeviceNo].Heating[2].Switch_ON_OFF <> "DB613_Komponent_State".Heating[0].Heating[2].Switch_ON_OFF OR
           "DB613_Komponent_State".Heating["DB613_Komponent_State".ReadDeviceNo].Heating[3].Switch_ON_OFF <> "DB613_Komponent_State".Heating[0].Heating[3].Switch_ON_OFF OR
           "DB613_Komponent_State".Heating["DB613_Komponent_State".ReadDeviceNo].Heating[4].Switch_ON_OFF <> "DB613_Komponent_State".Heating[0].Heating[4].Switch_ON_OFF OR
           "DB613_Komponent_State".Heating["DB613_Komponent_State".ReadDeviceNo].Heating[5].Switch_ON_OFF <> "DB613_Komponent_State".Heating[0].Heating[5].Switch_ON_OFF OR
           "DB613_Komponent_State".Heating["DB613_Komponent_State".ReadDeviceNo].Heating[6].Switch_ON_OFF <> "DB613_Komponent_State".Heating[0].Heating[6].Switch_ON_OFF OR
           "DB613_Komponent_State".Heating["DB613_Komponent_State".ReadDeviceNo].Heating[7].Switch_ON_OFF <> "DB613_Komponent_State".Heating[0].Heating[7].Switch_ON_OFF OR
           "DB613_Komponent_State".Heating["DB613_Komponent_State".ReadDeviceNo].Heating[8].Switch_ON_OFF <> "DB613_Komponent_State".Heating[0].Heating[8].Switch_ON_OFF
       THEN
           // copy the [0] switch to the selected switch
           "DB613_Komponent_State".Heating["DB613_Komponent_State".ReadDeviceNo].Heating[1].Switch_ON_OFF := "DB613_Komponent_State".Heating[0].Heating[1].Switch_ON_OFF;
           "DB613_Komponent_State".Heating["DB613_Komponent_State".ReadDeviceNo].Heating[2].Switch_ON_OFF := "DB613_Komponent_State".Heating[0].Heating[2].Switch_ON_OFF;
           "DB613_Komponent_State".Heating["DB613_Komponent_State".ReadDeviceNo].Heating[3].Switch_ON_OFF := "DB613_Komponent_State".Heating[0].Heating[3].Switch_ON_OFF;
           "DB613_Komponent_State".Heating["DB613_Komponent_State".ReadDeviceNo].Heating[4].Switch_ON_OFF := "DB613_Komponent_State".Heating[0].Heating[4].Switch_ON_OFF;
           "DB613_Komponent_State".Heating["DB613_Komponent_State".ReadDeviceNo].Heating[5].Switch_ON_OFF := "DB613_Komponent_State".Heating[0].Heating[5].Switch_ON_OFF;
           "DB613_Komponent_State".Heating["DB613_Komponent_State".ReadDeviceNo].Heating[6].Switch_ON_OFF := "DB613_Komponent_State".Heating[0].Heating[6].Switch_ON_OFF;
           "DB613_Komponent_State".Heating["DB613_Komponent_State".ReadDeviceNo].Heating[7].Switch_ON_OFF := "DB613_Komponent_State".Heating[0].Heating[7].Switch_ON_OFF;
           "DB613_Komponent_State".Heating["DB613_Komponent_State".ReadDeviceNo].Heating[8].Switch_ON_OFF := "DB613_Komponent_State".Heating[0].Heating[8].Switch_ON_OFF;
       ELSE
           // Read the status of the selected hydraulic
           "DB613_Komponent_State".Heating[0] := "DB613_Komponent_State".Heating["DB613_Komponent_State".ReadDeviceNo];
       END_IF;

   END_IF;


   // Write the nessesary information to the status area
   IF "DB613_Komponent_State".Write OR "DB608_PV_Metering".Write THEN
       // Write all prozess values
       "DB601_PV_Plunger".Component["DB613_Komponent_State".ReadDeviceNo] := "DB601_PV_Plunger".Component[0];
       "DB608_PV_Metering".Metering["DB613_Komponent_State".ReadDeviceNo].Flow := "DB608_PV_Metering".Metering[0].Flow;
       "DB608_PV_Metering".Metering["DB613_Komponent_State".ReadDeviceNo].Pressure := "DB608_PV_Metering".Metering[0].Pressure;
       "DB608_PV_Metering".Metering["DB613_Komponent_State".ReadDeviceNo].Temperature := "DB608_PV_Metering".Metering[0].Temperature;
       "DB608_PV_Metering".Metering["DB613_Komponent_State".ReadDeviceNo].Pre_Pressure := "DB608_PV_Metering".Metering[0].Pre_Pressure;
       "DB608_PV_Metering".Metering["DB613_Komponent_State".ReadDeviceNo].MixingRatio := "DB608_PV_Metering".Metering[0].MixingRatio;

       // + Temperierung    
       "DB608_PV_Metering".HeatexchangerHP["DB613_Komponent_State".ReadDeviceNo] := "DB608_PV_Metering".HeatexchangerHP[0];
       "DB608_PV_Metering".HeatexchangerLP["DB613_Komponent_State".ReadDeviceNo] := "DB608_PV_Metering".HeatexchangerLP[0];

       "DB608_PV_Metering".Heating["DB613_Komponent_State".ReadDeviceNo] := "DB608_PV_Metering".Heating[0];

       // Config values   
       "DB751_auxiliaryDriveMetering".FeedingPump["DB613_Komponent_State".ReadDeviceNo] := "DB751_auxiliaryDriveMetering".FeedingPump[0];
       "DB751_auxiliaryDriveMetering".EdgeFilter["DB613_Komponent_State".ReadDeviceNo] := "DB751_auxiliaryDriveMetering".EdgeFilter[0];
       "DB751_auxiliaryDriveMetering".HeatConverter["DB613_Komponent_State".ReadDeviceNo] := "DB751_auxiliaryDriveMetering".HeatConverter[0];
       "DB751_auxiliaryDriveMetering".HeatexchangerHP["DB613_Komponent_State".ReadDeviceNo] := "DB751_auxiliaryDriveMetering".HeatexchangerHP[0];
       "DB751_auxiliaryDriveMetering".HeatexchangerLP["DB613_Komponent_State".ReadDeviceNo] := "DB751_auxiliaryDriveMetering".HeatexchangerLP[0];
       "DB751_auxiliaryDriveMetering".FeedingPumpControler["DB613_Komponent_State".ReadDeviceNo] := "DB751_auxiliaryDriveMetering".FeedingPumpControler[0];

       "DB753_MeteringPump".Pump["DB613_Komponent_State".ReadDeviceNo] := "DB753_MeteringPump".Pump[0];
       "DB753_MeteringPump".HeatingController["DB613_Komponent_State".ReadDeviceNo] := "DB753_MeteringPump".HeatingController[0];
       "DB753_MeteringPump".Heating["DB613_Komponent_State".ReadDeviceNo] := "DB753_MeteringPump".Heating[0];

       //    "DB761_Cylinder_Manager".CylinderMan_Ma["DB613_Komponent_State".ReadWriteDeviceNo] := "DB761_Cylinder_Manager".CylinderMan_Ma[0];
       "DB762_Cylinder".Cylinder["DB613_Komponent_State".ReadDeviceNo] := "DB762_Cylinder".Cylinder[0];

       // Write special Flow values 
       "DB902_ConfFlow_PV".Flow["DB613_Komponent_State".ReadDeviceNo].controltime := "DB902_ConfFlow_PV".Flow[0].controltime;
       // Config Bits schieben
       // Feedimng Pump:
       "DB751_auxiliaryDriveMetering".FeedingPump[0].Config_Exist := "DB753_MeteringPump".Pump[0].WithFeedPump;
       "DB751_auxiliaryDriveMetering".FeedingPump["DB613_Komponent_State".ReadDeviceNo].Config_Exist := "DB751_auxiliaryDriveMetering".FeedingPump[0].Config_Exist;
       // EdgeFilter:
       "DB751_auxiliaryDriveMetering".EdgeFilter[0].Config_Exist := "DB753_MeteringPump".Pump[0].WithEdgeFilter;
       "DB751_auxiliaryDriveMetering".EdgeFilter["DB613_Komponent_State".ReadDeviceNo].Config_Exist := "DB751_auxiliaryDriveMetering".EdgeFilter[0].Config_Exist;
       //-----

   END_IF;

       "DB608_PV_Metering".Write := FALSE;
       "DB613_Komponent_State".Write := FALSE;

     // Show the actual values every time:
     "DB608_PV_Metering".Metering[0].Flow.PV_ActV := "DB608_PV_Metering".Metering["DB613_Komponent_State".ReadDeviceNo].Flow.PV_ActV;
     "DB608_PV_Metering".Metering[0].Pressure.PV_ActV := "DB608_PV_Metering".Metering["DB613_Komponent_State".ReadDeviceNo].Pressure.PV_ActV;
     "DB608_PV_Metering".Metering[0].Temperature.PV_ActV := "DB608_PV_Metering".Metering["DB613_Komponent_State".ReadDeviceNo].Temperature.PV_ActV;
     "DB608_PV_Metering".Metering[0].Pre_Pressure.PV_ActV := "DB608_PV_Metering".Metering["DB613_Komponent_State".ReadDeviceNo].Pre_Pressure.PV_ActV;
     "DB608_PV_Metering".Metering[0].MixingRatio.PV_ActV := "DB608_PV_Metering".Metering["DB613_Komponent_State".ReadDeviceNo].MixingRatio.PV_ActV;
     "DB608_PV_Metering".HeatexchangerHP[0].PV_ActV := "DB608_PV_Metering".HeatexchangerHP["DB613_Komponent_State".ReadDeviceNo].PV_ActV;
     "DB608_PV_Metering".HeatexchangerLP[0].PV_ActV := "DB608_PV_Metering".HeatexchangerLP["DB613_Komponent_State".ReadDeviceNo].PV_ActV;
     "DB608_PV_Metering".Heating[0].Heating[1].PV_ActV := "DB608_PV_Metering".Heating["DB613_Komponent_State".ReadDeviceNo].Heating[1].PV_ActV;
     "DB608_PV_Metering".Heating[0].Heating[2].PV_ActV := "DB608_PV_Metering".Heating["DB613_Komponent_State".ReadDeviceNo].Heating[2].PV_ActV;
     "DB608_PV_Metering".Heating[0].Heating[3].PV_ActV := "DB608_PV_Metering".Heating["DB613_Komponent_State".ReadDeviceNo].Heating[3].PV_ActV;
     "DB608_PV_Metering".Heating[0].Heating[4].PV_ActV := "DB608_PV_Metering".Heating["DB613_Komponent_State".ReadDeviceNo].Heating[4].PV_ActV;
     "DB608_PV_Metering".Heating[0].Heating[5].PV_ActV := "DB608_PV_Metering".Heating["DB613_Komponent_State".ReadDeviceNo].Heating[5].PV_ActV;
     "DB608_PV_Metering".Heating[0].Heating[6].PV_ActV := "DB608_PV_Metering".Heating["DB613_Komponent_State".ReadDeviceNo].Heating[6].PV_ActV;
     "DB608_PV_Metering".Heating[0].Heating[7].PV_ActV := "DB608_PV_Metering".Heating["DB613_Komponent_State".ReadDeviceNo].Heating[7].PV_ActV;
     "DB608_PV_Metering".Heating[0].Heating[8].PV_ActV := "DB608_PV_Metering".Heating["DB613_Komponent_State".ReadDeviceNo].Heating[8].PV_ActV;
END_FUNCTION

FUNCTION "FC5014_InterfaceMixinghead" : Void   // FC5014, SCL
{ S7_Optimized_Access := 'FALSE' }
VERSION : 0.1
   VAR_INPUT
      Enable : Bool;
   END_VAR
BEGIN

   // Read all values for the first selection
   IF ("DB614_MH_State".ReadDeviceNo <> "DB614_MH_State".ActualDeviceNo) OR "DB614_MH_State".Read THEN
       "DB614_MH_State".ActualDeviceNo := "DB614_MH_State".ReadDeviceNo;

       // Process values
       "DB604_PV_Mixinghead".Mixinghead[0] :="DB604_PV_Mixinghead".Mixinghead["DB614_MH_State".ReadDeviceNo];
       // Status
       "DB614_MH_State".MH_Status[0] := "DB614_MH_State".MH_Status["DB614_MH_State".ReadDeviceNo];
       // Sset values
       "DB704_MH_Value".Mixinghead[0] := "DB704_MH_Value".Mixinghead["DB614_MH_State".ReadDeviceNo];
       "DB704_MH_Value".MH_Inerting[0] := "DB704_MH_Value".MH_Inerting["DB614_MH_State".ReadDeviceNo];

       "DB614_MH_State".Read := FALSE;

   END_IF;

   // If not the mixinghead page was selectet don't save teh values   
   IF "TP-Bereichszeiger".Picturenumber.Bildnummer = 4 THEN
       IF NOT "DB123_MH_IO_Signals".MH[0].IN.MH_Manual_Mode = TRUE OR
           "DB619_State_MPart".Recirculation[1].Switch_Lowpressure = TRUE OR
           "DB619_State_MPart".Recirculation[1].Switch_Reduced = TRUE
       THEN
           "DB614_MH_State".MH_Status[0].Switch_Testshot_A_ON_OFF := FALSE;
           "DB614_MH_State".MH_Status[0].Switch_Testshot_B_ON_OFF := FALSE;
       END_IF;

       // If a status changed by operator copy this to the select number and do not read all status values
       IF "DB614_MH_State".MH_Status["DB614_MH_State".ReadDeviceNo].Switch_Service_ON_OFF <> "DB614_MH_State".MH_Status[0].Switch_Service_ON_OFF OR
           "DB614_MH_State".MH_Status["DB614_MH_State".ReadDeviceNo].Switch_HP_ON_OFF <> "DB614_MH_State".MH_Status[0].Switch_HP_ON_OFF OR
           "DB614_MH_State".MH_Status["DB614_MH_State".ReadDeviceNo].QPB_Values_selected <> "DB614_MH_State".MH_Status[0].QPB_Values_selected OR
           "DB614_MH_State".MH_Status["DB614_MH_State".ReadDeviceNo].Switch_Testshot_A_ON_OFF <> "DB614_MH_State".MH_Status[0].Switch_Testshot_A_ON_OFF OR
           "DB614_MH_State".MH_Status["DB614_MH_State".ReadDeviceNo].Switch_Testshot_B_ON_OFF <> "DB614_MH_State".MH_Status[0].Switch_Testshot_B_ON_OFF
       THEN
           "DB614_MH_State".MH_Status["DB614_MH_State".ReadDeviceNo].Switch_Service_ON_OFF := "DB614_MH_State".MH_Status[0].Switch_Service_ON_OFF;
           "DB614_MH_State".MH_Status["DB614_MH_State".ReadDeviceNo].Switch_HP_ON_OFF := "DB614_MH_State".MH_Status[0].Switch_HP_ON_OFF;
           "DB614_MH_State".MH_Status["DB614_MH_State".ReadDeviceNo].QPB_Values_selected := "DB614_MH_State".MH_Status[0].QPB_Values_selected;
           "DB614_MH_State".MH_Status["DB614_MH_State".ReadDeviceNo].Switch_Testshot_A_ON_OFF := "DB614_MH_State".MH_Status[0].Switch_Testshot_A_ON_OFF;
           "DB614_MH_State".MH_Status["DB614_MH_State".ReadDeviceNo].Switch_Testshot_B_ON_OFF := "DB614_MH_State".MH_Status[0].Switch_Testshot_B_ON_OFF;
       ELSE
           "DB614_MH_State".MH_Status[0] := "DB614_MH_State".MH_Status["DB614_MH_State".ReadDeviceNo];
       END_IF;

       // If a status for the cleaning pisteon changed by operator copy this to the select number and do not read all status values
       IF "DB614_MH_State".MH_CleaningPiston["DB614_MH_State".ReadDeviceNo].Switch_CP_Forward <> "DB614_MH_State".MH_CleaningPiston[0].Switch_CP_Forward
       THEN
           "DB614_MH_State".MH_CleaningPiston["DB614_MH_State".ReadDeviceNo].Switch_CP_Forward := "DB614_MH_State".MH_CleaningPiston[0].Switch_CP_Forward;
       ELSE
           "DB614_MH_State".MH_CleaningPiston[0] := "DB614_MH_State".MH_CleaningPiston["DB614_MH_State".ReadDeviceNo];
       END_IF;

       // If a status for the mixinghead look system changed by operator copy this to the select number and do not read all status values
       IF "DB614_MH_State".MH_Lock["DB614_MH_State".ReadDeviceNo].Switch_MH_Lock_ON_OFF <> "DB614_MH_State".MH_Lock[0].Switch_MH_Lock_ON_OFF
       THEN
           "DB614_MH_State".MH_Lock["DB614_MH_State".ReadDeviceNo].Switch_MH_Lock_ON_OFF := "DB614_MH_State".MH_Lock[0].Switch_MH_Lock_ON_OFF;
       ELSE
           "DB614_MH_State".MH_Lock[0] := "DB614_MH_State".MH_Lock["DB614_MH_State".ReadDeviceNo];
       END_IF;